   "DB302_HMI_Faults_Carrier71_Faults_1" : Int = PLC DB302_HMI_Faults.Carrier71_Faults_1 AT %DB1.DBW0, 1 s
   "DB302_HMI_Faults_Carrier71_Faults_2" : Int = PLC DB302_HMI_Faults.Carrier71_Faults_2 AT %DB1.DBW0, 1 s
   "DB302_HMI_Faults_Carrier71_Faults_3" : Int = PLC DB302_HMI_Faults.Carrier71_Faults_3 AT %DB1.DBW0, 1 s
   "DB302_HMI_Faults_Carrier72_Faults_0" : Int = PLC DB302_HMI_Faults.Carrier72_Faults_0 AT %DB1.DBW0, 1 s
   "DB302_HMI_Faults_Carrier72_Faults_1" : Int = PLC DB302_HMI_Faults.Carrier72_Faults_1 AT %DB1.DBW0, 1 s
   "DB302_HMI_Faults_Carrier72_Faults_2" : Int = PLC DB302_HMI_Faults.Carrier72_Faults_2 AT %DB1.DBW0, 1 s
   "DB302_HMI_Faults_Carrier72_Faults_3" : Int = PLC DB302_HMI_Faults.Carrier72_Faults_3 AT %DB1.DBW0, 1 s
   "DB302_HMI_Faults_Carrier73_Faults_0" : Int = PLC DB302_HMI_Faults.Carrier73_Faults_0 AT %DB1.DBW0, 1 s
   "DB302_HMI_Faults_Carrier73_Faults_1" : Int = PLC DB302_HMI_Faults.Carrier73_Faults_1 AT %DB1.DBW0, 1 s
   "DB302_HMI_Faults_Carrier73_Faults_2" : Int = PLC DB302_HMI_Faults.Carrier73_Faults_2 AT %DB1.DBW0, 1 s
   "DB302_HMI_Faults_Carrier73_Faults_3" : Int = PLC DB302_HMI_Faults.Carrier73_Faults_3 AT %DB1.DBW0, 1 s
   "DB302_HMI_Faults_Carrier74_Faults_0" : Int = PLC DB302_HMI_Faults.Carrier74_Faults_0 AT %DB1.DBW0, 1 s
   "DB302_HMI_Faults_Carrier74_Faults_1" : Int = PLC DB302_HMI_Faults.Carrier74_Faults_1 AT %DB1.DBW0, 1 s
   "DB302_HMI_Faults_Carrier74_Faults_2" : Int = PLC DB302_HMI_Faults.Carrier74_Faults_2 AT %DB1.DBW0, 1 s
   "DB302_HMI_Faults_Carrier74_Faults_3" : Int = PLC DB302_HMI_Faults.Carrier74_Faults_3 AT %DB1.DBW0, 1 s
   "DB302_HMI_Faults_Carrier75_Faults_0" : Int = PLC DB302_HMI_Faults.Carrier75_Faults_0 AT %DB1.DBW0, 1 s
   "DB302_HMI_Faults_Carrier75_Faults_1" : Int = PLC DB302_HMI_Faults.Carrier75_Faults_1 AT %DB1.DBW0, 1 s
   "DB302_HMI_Faults_Carrier75_Faults_2" : Int = PLC DB302_HMI_Faults.Carrier75_Faults_2 AT %DB1.DBW0, 1 s
   "DB302_HMI_Faults_Carrier75_Faults_3" : Int = PLC DB302_HMI_Faults.Carrier75_Faults_3 AT %DB1.DBW0, 1 s
   "DB302_HMI_Faults_Carrier76_Faults_0" : Int = PLC DB302_HMI_Faults.Carrier76_Faults_0 AT %DB1.DBW0, 1 s
   "DB302_HMI_Faults_Carrier76_Faults_1" : Int = PLC DB302_HMI_Faults.Carrier76_Faults_1 AT %DB1.DBW0, 1 s
   "DB302_HMI_Faults_Carrier76_Faults_2" : Int = PLC DB302_HMI_Faults.Carrier76_Faults_2 AT %DB1.DBW0, 1 s
   "DB302_HMI_Faults_Carrier76_Faults_3" : Int = PLC DB302_HMI_Faults.Carrier76_Faults_3 AT %DB1.DBW0, 1 s
   "DB302_HMI_Faults_Carrier77_Faults_0" : Int = PLC DB302_HMI_Faults.Carrier77_Faults_0 AT %DB1.DBW0, 1 s
   "DB302_HMI_Faults_Carrier77_Faults_1" : Int = PLC DB302_HMI_Faults.Carrier77_Faults_1 AT %DB1.DBW0, 1 s
   "DB302_HMI_Faults_Carrier77_Faults_2" : Int = PLC DB302_HMI_Faults.Carrier77_Faults_2 AT %DB1.DBW0, 1 s
   "DB302_HMI_Faults_Carrier77_Faults_3" : Int = PLC DB302_HMI_Faults.Carrier77_Faults_3 AT %DB1.DBW0, 1 s
   "DB302_HMI_Faults_Carrier78_Faults_0" : Int = PLC DB302_HMI_Faults.Carrier78_Faults_0 AT %DB1.DBW0, 1 s
   "DB302_HMI_Faults_Carrier78_Faults_1" : Int = PLC DB302_HMI_Faults.Carrier78_Faults_1 AT %DB1.DBW0, 1 s
   "DB302_HMI_Faults_Carrier78_Faults_2" : Int = PLC DB302_HMI_Faults.Carrier78_Faults_2 AT %DB1.DBW0, 1 s
   "DB302_HMI_Faults_Carrier78_Faults_3" : Int = PLC DB302_HMI_Faults.Carrier78_Faults_3 AT %DB1.DBW0, 1 s
   "DB302_HMI_Faults_Carrier79_Faults_0" : Int = PLC DB302_HMI_Faults.Carrier79_Faults_0 AT %DB1.DBW0, 1 s
   "DB302_HMI_Faults_Carrier79_Faults_1" : Int = PLC DB302_HMI_Faults.Carrier79_Faults_1 AT %DB1.DBW0, 1 s
   "DB302_HMI_Faults_Carrier79_Faults_2" : Int = PLC DB302_HMI_Faults.Carrier79_Faults_2 AT %DB1.DBW0, 1 s
   "DB302_HMI_Faults_Carrier79_Faults_3" : Int = PLC DB302_HMI_Faults.Carrier79_Faults_3 AT %DB1.DBW0, 1 s
   "DB302_HMI_Faults_Carrier8_Faults_0" : Int = PLC DB302_HMI_Faults.Carrier8_Faults_0 AT %DB1.DBW0, 1 s
   "DB302_HMI_Faults_Carrier8_Faults_1" : Int = PLC DB302_HMI_Faults.Carrier8_Faults_1 AT %DB1.DBW0, 1 s
   "DB302_HMI_Faults_Carrier8_Faults_2" : Int = PLC DB302_HMI_Faults.Carrier8_Faults_2 AT %DB1.DBW0, 1 s
   "DB302_HMI_Faults_Carrier8_Faults_3" : Int = PLC DB302_HMI_Faults.Carrier8_Faults_3 AT %DB1.DBW0, 1 s
   "DB302_HMI_Faults_Carrier80_Faults_0" : Int = PLC DB302_HMI_Faults.Carrier80_Faults_0 AT %DB1.DBW0, 1 s
   "DB302_HMI_Faults_Carrier80_Faults_1" : Int = PLC DB302_HMI_Faults.Carrier80_Faults_1 AT %DB1.DBW0, 1 s
   "DB302_HMI_Faults_Carrier80_Faults_2" : Int = PLC DB302_HMI_Faults.Carrier80_Faults_2 AT %DB1.DBW0, 1 s
   "DB302_HMI_Faults_Carrier80_Faults_3" : Int = PLC DB302_HMI_Faults.Carrier80_Faults_3 AT %DB1.DBW0, 1 s
   "DB302_HMI_Faults_Carrier81_Faults_0" : Int = PLC DB302_HMI_Faults.Carrier81_Faults_0 AT %DB1.DBW0, 1 s
   "DB302_HMI_Faults_Carrier81_Faults_1" : Int = PLC DB302_HMI_Faults.Carrier81_Faults_1 AT %DB1.DBW0, 1 s
   "DB302_HMI_Faults_Carrier81_Faults_2" : Int = PLC DB302_HMI_Faults.Carrier81_Faults_2 AT %DB1.DBW0, 1 s
   "DB302_HMI_Faults_Carrier81_Faults_3" : Int = PLC DB302_HMI_Faults.Carrier81_Faults_3 AT %DB1.DBW0, 1 s
   "DB302_HMI_Faults_Carrier82_Faults_0" : Int = PLC DB302_HMI_Faults.Carrier82_Faults_0 AT %DB1.DBW0, 1 s
   "DB302_HMI_Faults_Carrier82_Faults_1" : Int = PLC DB302_HMI_Faults.Carrier82_Faults_1 AT %DB1.DBW0, 1 s
   "DB302_HMI_Faults_Carrier82_Faults_2" : Int = PLC DB302_HMI_Faults.Carrier82_Faults_2 AT %DB1.DBW0, 1 s
   "DB302_HMI_Faults_Carrier82_Faults_3" : Int = PLC DB302_HMI_Faults.Carrier82_Faults_3 AT %DB1.DBW0, 1 s
   "DB302_HMI_Faults_Carrier9_Faults_0" : Int = PLC DB302_HMI_Faults.Carrier9_Faults_0 AT %DB1.DBW0, 1 s
   "DB302_HMI_Faults_Carrier9_Faults_1" : Int = PLC DB302_HMI_Faults.Carrier9_Faults_1 AT %DB1.DBW0, 1 s
   "DB302_HMI_Faults_Carrier9_Faults_2" : Int = PLC DB302_HMI_Faults.Carrier9_Faults_2 AT %DB1.DBW0, 1 s
   "DB302_HMI_Faults_Carrier9_Faults_3" : Int = PLC DB302_HMI_Faults.Carrier9_Faults_3 AT %DB1.DBW0, 1 s
   "DB401_HMI_Status_ZoneStatus.AccumZoneSpacing" : Word = PLC DB401_HMI_Status.ZoneStatus.AccumZoneSpacing, 1 s
   "DB401_HMI_Status_ZoneStatus.NextZoneNumber" : Int = PLC DB401_HMI_Status.ZoneStatus.NextZoneNumber, 1 s
   "DB401_HMI_Status_ZoneStatus.ProductionZoneSpacing" : Word = PLC DB401_HMI_Status.ZoneStatus.ProductionZoneSpacing, 1 s
   "DB401_HMI_Status_ZoneStatus.SpeedZone" : Bool = PLC DB401_HMI_Status.ZoneStatus.SpeedZone, 1 s
   "DB401_HMI_Status_ZoneStatus.SpeedZoneEndPos" : DWord = PLC DB401_HMI_Status.ZoneStatus.SpeedZoneEndPos, 1 s
   "DB401_HMI_Status_ZoneStatus.SpeedZoneStartPos" : DWord = PLC DB401_HMI_Status.ZoneStatus.SpeedZoneStartPos, 1 s
   "DB401_HMI_Status_ZoneStatus.ZoneEndPosition" : DWord = PLC DB401_HMI_Status.ZoneStatus.ZoneEndPosition, 1 s
   "DB401_HMI_Status_ZoneStatus.ZoneFull" : Bool = PLC DB401_HMI_Status.ZoneStatus.ZoneFull, 1 s
   "DB401_HMI_Status_ZoneStatus.ZoneIndex" : Int = PLC DB401_HMI_Status.ZoneStatus.ZoneIndex, 1 s
   "DB401_HMI_Status_ZoneStatus.ZoneStartPosition" : DWord = PLC DB401_HMI_Status.ZoneStatus.ZoneStartPosition, 1 s
   "DB401_HMI_Status_ZoneStatus.ZoneType" : String[254] = PLC DB401_HMI_Status.ZoneStatus.ZoneType, 1 s
   "DB401_HMI_Status_CarrierFaultCode" : Int = PLC DB401_HMI_Status.Status.CarrierFaultCode, 1 s
   "EMS_Zone[31]" : UDT_ZoneStructure = PLC EMS.Zone[31] AT %DB8.DBX31020.0, 1 s
   "EMS_Zone[32]" : UDT_ZoneStructure = PLC EMS.Zone[32] AT %DB8.DBX31020.0, 1 s
   "EMS_Zone[33]" : UDT_ZoneStructure = PLC EMS.Zone[33] AT %DB1.DBW0, 1 s
   "EMS_Zone[34]" : UDT_ZoneStructure = PLC EMS.Zone[34] AT %DB1.DBW0, 1 s
   "EMS_Zone[35]" : UDT_ZoneStructure = PLC EMS.Zone[35] AT %DB1.DBW0, 1 s
   "EMS_Zone[36]" : UDT_ZoneStructure = PLC EMS.Zone[36] AT %DB1.DBW0, 1 s
   "EMS_Zone[37]" : UDT_ZoneStructure = PLC EMS.Zone[37] AT %DB1.DBW0, 1 s
   "EMS_Zone[38]" : UDT_ZoneStructure = PLC EMS.Zone[38] AT %DB1.DBW0, 1 s
   "EMS_Zone[39]" : UDT_ZoneStructure = PLC EMS.Zone[39] AT %DB1.DBW0, 1 s
   "EMS_Zone[4]" : UDT_ZoneStructure = PLC EMS.Zone[4] AT %DB8.DBX4136.0, 1 s
   "EMS_Zone[40]" : UDT_ZoneStructure = PLC EMS.Zone[40] AT %DB1.DBW0, 1 s
   "EMS_Zone[41]" : UDT_ZoneStructure = PLC EMS.Zone[41] AT %DB1.DBW0, 1 s
   "EMS_Zone[42]" : UDT_ZoneStructure = PLC EMS.Zone[42] AT %DB1.DBW0, 1 s
   "EMS_Zone[43]" : UDT_ZoneStructure = PLC EMS.Zone[43] AT %DB1.DBW0, 1 s
   "EMS_Zone[44]" : UDT_ZoneStructure = PLC EMS.Zone[44] AT %DB1.DBW0, 1 s
   "EMS_Zone[45]" : UDT_ZoneStructure = PLC EMS.Zone[45] AT %DB1.DBW0, 1 s
   "EMS_Zone[46]" : UDT_ZoneStructure = PLC EMS.Zone[46] AT %DB1.DBW0, 1 s
   "EMS_Zone[47]" : UDT_ZoneStructure = PLC EMS.Zone[47] AT %DB1.DBW0, 1 s
   "EMS_Zone[48]" : UDT_ZoneStructure = PLC EMS.Zone[48] AT %DB1.DBW0, 1 s
   "EMS_Zone[49]" : UDT_ZoneStructure = PLC EMS.Zone[49] AT %DB1.DBW0, 1 s
   "EMS_Zone[5]" : UDT_ZoneStructure = PLC EMS.Zone[5] AT %DB8.DBX5170.0, 1 s
   "EMS_Zone[50]" : UDT_ZoneStructure = PLC EMS.Zone[50] AT %DB1.DBW0, 1 s
   "EMS_Zone[51]" : UDT_ZoneStructure = PLC EMS.Zone[51] AT %DB1.DBW0, 1 s
   "EMS_Zone[52]" : UDT_ZoneStructure = PLC EMS.Zone[52] AT %DB8.DBX31020.0, 1 s
   "EMS_Zone[53]" : UDT_ZoneStructure = PLC EMS.Zone[53] AT %DB1.DBW0, 1 s
   "EMS_Zone[54]" : UDT_ZoneStructure = PLC EMS.Zone[54] AT %DB1.DBW0, 1 s
   "EMS_Zone[55]" : UDT_ZoneStructure = PLC EMS.Zone[55] AT %DB1.DBW0, 1 s
   "EMS_Zone[56]" : UDT_ZoneStructure = PLC EMS.Zone[56] AT %DB1.DBW0, 1 s
   "EMS_Zone[57]" : UDT_ZoneStructure = PLC EMS.Zone[57] AT %DB1.DBW0, 1 s
   "EMS_Zone[58]" : UDT_ZoneStructure = PLC EMS.Zone[58] AT %DB8.DBX31020.0, 1 s
   "EMS_Zone[59]" : UDT_ZoneStructure = PLC EMS.Zone[59] AT %DB1.DBW0, 1 s
   "EMS_Zone[6]" : UDT_ZoneStructure = PLC EMS.Zone[6] AT %DB8.DBX6204.0, 1 s
   "EMS_Zone[60]" : UDT_ZoneStructure = PLC EMS.Zone[60] AT %DB1.DBW0, 1 s
   "EMS_Zone[61]" : UDT_ZoneStructure = PLC EMS.Zone[61] AT %DB1.DBW0, 1 s
   "EMS_Zone[62]" : UDT_ZoneStructure = PLC EMS.Zone[62] AT %DB1.DBW0, 1 s
   "EMS_Zone[63]" : UDT_ZoneStructure = PLC EMS.Zone[63] AT %DB1.DBW0, 1 s
   "DB401_HMI_Status_ZoneStatus.PrevZoneNumber" : Int = PLC DB401_HMI_Status.ZoneStatus.PrevZoneNumber, 1 s
   "Mask_Carrier_Faults_LT" : Bool = PLC DB401_HMI_Status.Status.MaskCarrierFaultsLT AT %DB1.DBX0.0, 1 s
   "Reset_Mask_Carrier_Faults_PB" : Bool = PLC DB401_HMI_Status.Status.ResetMaskCarrierFaultsPB AT %DB1.DBX0.0, 1 s
   "Set_Mask_Carrier_Faults_PB" : Bool = PLC DB401_HMI_Status.Status.SetMaskCarrierFaultsPB AT %DB1.DBX0.0, 1 s
   "HMI_Carrier_CurrentArea" : String[2] = PLC DB401_HMI_Status.Status.Area AT %DB1.DBW0, 1 s

HMI tags "SDC"
   "Clock_1Hz" : Bool = PLC Clock_1Hz AT %M0.5, 500 ms   // Zyklusflanke 1Hz / Cycle flag 1Hz
   "SDC\_EDIT" : Int, internal
   "SDC\_EDIT_BIT" : Bool, internal
   "SDC\_open_EMS_Stat" : Bool, internal
      on ChangeValue: ActivateScreen("711_CARRIER_STATUS", 0)
   "SDC\_open_Section_Para" : Bool, internal
      on ChangeValue: ActivateScreen("708_ZONE_STATUS", 0)
   "HMI_EMS_Nr" : Int = PLC HMI_EMS_Nr AT %MW30, 1 s
   "SDC\_TS_Nr" : Int, internal
      on ChangeValue: "SDC_TS_PARAMETER"(); "SDC_TS_REFERENCE"("SDC\_TS_Nr")
   "SDC\_intern_Bildnummer" : Int AT %DB1.DBX0.0
   "DB_SDC_GLOBAL_M.SDC_ER_Reset" : Bool = PLC DB_SDC_GLOBAL.M.SDC_ER_Reset AT %DB3700.DBX600.4, 1 s
   "SDC\_intern_MELDUNGEN" : Int, internal
   "SDC\_Pos_sichtbar" : Bool AT %DB1.DBX4.0
   "AlwaysTRUE" : Bool = PLC AlwaysTRUE AT %M1.2, 500 ms
   "AlwaysFALSE" : Bool = PLC AlwaysFALSE AT %M1.3, 500 ms
   "HMI_Zone_Nr" : Int = PLC HMI_Zone_Nr AT %MW102, 1 s
   "HMI_Status_G120D_Control" : Word = PLC DB401_HMI_Status.Drive.G120D_CONTROL AT %DB1.DBW0, 1 s
   "HMI_Status_G120D_Status" : Word = PLC DB401_HMI_Status.Drive.G120D_STATUS AT %DB1.DBW0, 1 s
   "HMI_Status_Slot2_Inputs" : Byte = PLC DB401_HMI_Status.IO.Carrier_Slot02_Inputs AT %DB1.DBW0, 1 s
   "HMI_Status_Slot3_Outputs" : Byte = PLC DB401_HMI_Status.IO.Carrier_Slot03_Outputs AT %DB1.DBW0, 1 s
   "HMI_Status_Slot4_Inputs" : Word = PLC DB401_HMI_Status.IO.Carrier_Slot04_Inputs AT %DB1.DBW0, 1 s
   "HMI_Status_Slot5_Outputs" : Word = PLC DB401_HMI_Status.IO.Carrier_Slot05_Outputs AT %DB1.DBW0, 1 s
   "HMI_Carrier_Comm_Fault" : Bool = PLC DB401_HMI_Status.Status.CommFlt AT %DB1.DBW0, 1 s
   "HMI_Carrier_Faulted" : Bool = PLC DB401_HMI_Status.Status.Faulted AT %DB1.DBW0, 1 s
   "HMI_Carrier_Auto" : Bool = PLC DB401_HMI_Status.Status.AutoMode AT %DB1.DBW0, 1 s
   "HMI_Carrier_Manual" : Bool = PLC DB401_HMI_Status.Status.ManualMode AT %DB1.DBW0, 1 s
   "HMI_Carrier_RunningFwd" : Bool = PLC DB401_HMI_Status.Status.RunningFWD AT %DB1.DBW0, 1 s
   "HMI_Carrier_RunningRev" : Bool = PLC DB401_HMI_Status.Status.RunningREV AT %DB1.DBW0, 1 s
   "HMI_Carrier_HoldPBPressed" : Bool = PLC DB401_HMI_Status.Status.ProductionHoldPB_Status AT %DB1.DBW0, 1 s
   "HMI_Carrier_DriveFwdCommand" : Bool = PLC DB401_HMI_Status.Status.DriveFwdCMD AT %DB1.DBW0, 1 s
   "HMI_Carrier_DriveCmdSpeed" : Word = PLC DB401_HMI_Status.Status.DriveCmdSpeed AT %DB1.DBW0, 1 s
   "HMI_Carrier_CurrentPosition" : DWord = PLC DB401_HMI_Status.Status.CarrierPosition AT %DB1.DBW0, 1 s
   "HMI_Carrier_ActualSpeed" : Word = PLC DB401_HMI_Status.Status.ActualSpeed AT %DB1.DBW0, 1 s
   "HMI_Carrier_NextCarrierNumber" : Word = PLC DB401_HMI_Status.Status.NextCarrierNum AT %DB1.DBW0, 1 s
   "HMI_Carrier_CurrentZone" : Int = PLC DB401_HMI_Status.Status.Zone AT %DB1.DBW0, 1 s
   "HMI_Carrier_AtCommandPosition" : Bool = PLC DB401_HMI_Status.Status.AtCmdPos AT %DB1.DBW0, 1 s
   "HMI_Carrier_NextStopPosition" : DWord = PLC DB401_HMI_Status.Status.NextStopPosition AT %DB1.DBW0, 1 s
   "HMI_Carrier_DriveCommFault" : Bool = PLC DB401_HMI_Status.Status.DriveCommFault AT %DB1.DBW0, 1 s
   "HMI_Carrier_EncoderCommFault" : Bool = PLC DB401_HMI_Status.Status.EncoderCommFault AT %DB1.DBW0, 1 s
   "HMI_Carrier_HMICommFault" : Bool = PLC DB401_HMI_Status.Status.HMICommFault AT %DB1.DBW0, 1 s

HMI tags "DB_SDC_EMS_TS_HMI"
   "DB_SDC_EMS_TS_1_HMI_SEK[88].EMS[1]" : UDT_SDC_EMS_TS_STAT_HMI = PLC DB_SDC_EMS_TS_1_HMI.SEK[88].EMS[1] AT %DB3810.DBX15680.0, 1 s
   "DB_SDC_EMS_TS_1_HMI_SEK[89].EMS[1]" : UDT_SDC_EMS_TS_STAT_HMI = PLC DB_SDC_EMS_TS_1_HMI.SEK[89].EMS[1] AT %DB3810.DBX15860.0, 1 s
   "DB_SDC_EMS_TS_1_HMI_SEK[90].EMS[1]" : UDT_SDC_EMS_TS_STAT_HMI = PLC DB_SDC_EMS_TS_1_HMI.SEK[90].EMS[1] AT %DB3810.DBX16040.0, 1 s
   "DB_SDC_EMS_TS_1_HMI_SEK[91].EMS[1]" : UDT_SDC_EMS_TS_STAT_HMI = PLC DB_SDC_EMS_TS_1_HMI.SEK[91].EMS[1] AT %DB3810.DBX16220.0, 1 s
   "DB_SDC_EMS_TS_1_HMI_SEK[92].EMS[1]" : UDT_SDC_EMS_TS_STAT_HMI = PLC DB_SDC_EMS_TS_1_HMI.SEK[92].EMS[1] AT %DB3810.DBX16400.0, 1 s
   "DB_SDC_EMS_TS_1_HMI_SEK[93].EMS[1]" : UDT_SDC_EMS_TS_STAT_HMI = PLC DB_SDC_EMS_TS_1_HMI.SEK[93].EMS[1] AT %DB3810.DBX16580.0, 1 s
   "DB_SDC_EMS_TS_1_HMI_SEK[94].EMS[1]" : UDT_SDC_EMS_TS_STAT_HMI = PLC DB_SDC_EMS_TS_1_HMI.SEK[94].EMS[1] AT %DB3810.DBX16760.0, 1 s
   "DB_SDC_EMS_TS_1_HMI_SEK[95].EMS[1]" : UDT_SDC_EMS_TS_STAT_HMI = PLC DB_SDC_EMS_TS_1_HMI.SEK[95].EMS[1] AT %DB3810.DBX16940.0, 1 s
   "DB_SDC_EMS_TS_1_HMI_SEK[96].EMS[1]" : UDT_SDC_EMS_TS_STAT_HMI = PLC DB_SDC_EMS_TS_1_HMI.SEK[96].EMS[1] AT %DB3810.DBX17120.0, 1 s
   "DB_SDC_EMS_TS_1_HMI_SEK[100].EMS[1]" : UDT_SDC_EMS_TS_STAT_HMI = PLC DB_SDC_EMS_TS_1_HMI.SEK[100].EMS[1] AT %DB3810.DBX17840.0, 1 s
   "DB_SDC_EMS_TS_1_HMI_SEK[101].EMS[1]" : UDT_SDC_EMS_TS_STAT_HMI = PLC DB_SDC_EMS_TS_1_HMI.SEK[101].EMS[1] AT %DB3810.DBX18020.0, 1 s
   "DB_SDC_EMS_TS_1_HMI_SEK[102].EMS[1]" : UDT_SDC_EMS_TS_STAT_HMI = PLC DB_SDC_EMS_TS_1_HMI.SEK[102].EMS[1] AT %DB3810.DBX18200.0, 1 s
   "DB_SDC_EMS_TS_1_HMI_SEK[103].EMS[1]" : UDT_SDC_EMS_TS_STAT_HMI = PLC DB_SDC_EMS_TS_1_HMI.SEK[103].EMS[1] AT %DB3810.DBX18380.0, 1 s
   "DB_SDC_EMS_TS_1_HMI_SEK[104].EMS[1]" : UDT_SDC_EMS_TS_STAT_HMI = PLC DB_SDC_EMS_TS_1_HMI.SEK[104].EMS[1] AT %DB3810.DBX18560.0, 1 s
   "DB_SDC_EMS_TS_1_HMI_SEK[105].EMS[1]" : UDT_SDC_EMS_TS_STAT_HMI = PLC DB_SDC_EMS_TS_1_HMI.SEK[105].EMS[1] AT %DB3810.DBX18740.0, 1 s
   "DB_SDC_EMS_TS_1_HMI_SEK[106].EMS[1]" : UDT_SDC_EMS_TS_STAT_HMI = PLC DB_SDC_EMS_TS_1_HMI.SEK[106].EMS[1] AT %DB3810.DBX18920.0, 1 s
   "DB_SDC_EMS_TS_1_HMI_SEK[107].EMS[1]" : UDT_SDC_EMS_TS_STAT_HMI = PLC DB_SDC_EMS_TS_1_HMI.SEK[107].EMS[1] AT %DB3810.DBX19100.0, 1 s
   "DB_SDC_EMS_TS_1_HMI_SEK[108].EMS[1]" : UDT_SDC_EMS_TS_STAT_HMI = PLC DB_SDC_EMS_TS_1_HMI.SEK[108].EMS[1] AT %DB3810.DBX19280.0, 1 s
   "DB_SDC_EMS_TS_1_HMI_SEK[109].EMS[1]" : UDT_SDC_EMS_TS_STAT_HMI = PLC DB_SDC_EMS_TS_1_HMI.SEK[109].EMS[1] AT %DB3810.DBX19460.0, 1 s
   "DB_SDC_EMS_TS_1_HMI_SEK[110].EMS[1]" : UDT_SDC_EMS_TS_STAT_HMI = PLC DB_SDC_EMS_TS_1_HMI.SEK[110].EMS[1] AT %DB3810.DBX19640.0, 1 s
   "DB_SDC_EMS_TS_1_HMI_SEK[111].EMS[1]" : UDT_SDC_EMS_TS_STAT_HMI = PLC DB_SDC_EMS_TS_1_HMI.SEK[111].EMS[1] AT %DB3810.DBX19820.0, 1 s
   "DB_SDC_EMS_TS_1_HMI_SEK[120].EMS[1]" : UDT_SDC_EMS_TS_STAT_HMI = PLC DB_SDC_EMS_TS_1_HMI.SEK[120].EMS[1] AT %DB3810.DBX21440.0, 1 s
   "DB_SDC_EMS_TS_1_HMI_SEK[121].EMS[1]" : UDT_SDC_EMS_TS_STAT_HMI = PLC DB_SDC_EMS_TS_1_HMI.SEK[121].EMS[1] AT %DB3810.DBX21620.0, 1 s
   "DB_SDC_EMS_TS_1_HMI_SEK[126].EMS[1]" : UDT_SDC_EMS_TS_STAT_HMI = PLC DB_SDC_EMS_TS_1_HMI.SEK[126].EMS[1] AT %DB3810.DBX22520.0, 1 s
   "DB_SDC_EMS_TS_1_HMI_SEK[125].EMS[1]" : UDT_SDC_EMS_TS_STAT_HMI = PLC DB_SDC_EMS_TS_1_HMI.SEK[125].EMS[1] AT %DB3810.DBX22340.0, 1 s
   "DB_SDC_EMS_TS_1_HMI_SEK[122].EMS[1]" : UDT_SDC_EMS_TS_STAT_HMI = PLC DB_SDC_EMS_TS_1_HMI.SEK[122].EMS[1] AT %DB3810.DBX21800.0, 1 s
   "DB_SDC_EMS_TS_1_HMI_SEK[123].EMS[1]" : UDT_SDC_EMS_TS_STAT_HMI = PLC DB_SDC_EMS_TS_1_HMI.SEK[123].EMS[1] AT %DB3810.DBX21980.0, 1 s
   "DB_SDC_EMS_TS_1_HMI_SEK[124].EMS[1]" : UDT_SDC_EMS_TS_STAT_HMI = PLC DB_SDC_EMS_TS_1_HMI.SEK[124].EMS[1] AT %DB3810.DBX22160.0, 1 s
   "DB_SDC_EMS_TS_1_HMI_SEK[127].EMS[1]" : UDT_SDC_EMS_TS_STAT_HMI = PLC DB_SDC_EMS_TS_1_HMI.SEK[127].EMS[1] AT %DB3810.DBX22700.0, 1 s
   "DB_SDC_EMS_TS_1_HMI_SEK[128].EMS[1]" : UDT_SDC_EMS_TS_STAT_HMI = PLC DB_SDC_EMS_TS_1_HMI.SEK[128].EMS[1] AT %DB3810.DBX22880.0, 1 s
   "DB_SDC_EMS_TS_1_HMI_SEK[129].EMS[1]" : UDT_SDC_EMS_TS_STAT_HMI = PLC DB_SDC_EMS_TS_1_HMI.SEK[129].EMS[1] AT %DB3810.DBX23060.0, 1 s
   "DB_SDC_EMS_TS_1_HMI_SEK[130].EMS[1]" : UDT_SDC_EMS_TS_STAT_HMI = PLC DB_SDC_EMS_TS_1_HMI.SEK[130].EMS[1] AT %DB3810.DBX23240.0, 1 s
   "DB_SDC_EMS_TS_1_HMI_SEK[131].EMS[1]" : UDT_SDC_EMS_TS_STAT_HMI = PLC DB_SDC_EMS_TS_1_HMI.SEK[131].EMS[1] AT %DB3810.DBX23420.0, 1 s
   "DB_SDC_EMS_TS_1_HMI_SEK[132].EMS[1]" : UDT_SDC_EMS_TS_STAT_HMI = PLC DB_SDC_EMS_TS_1_HMI.SEK[132].EMS[1] AT %DB3810.DBX23600.0, 1 s
   "DB_SDC_EMS_TS_1_HMI_SEK[140].EMS[1]" : UDT_SDC_EMS_TS_STAT_HMI = PLC DB_SDC_EMS_TS_1_HMI.SEK[140].EMS[1] AT %DB3810.DBX25040.0, 1 s
   "DB_SDC_EMS_TS_1_HMI_SEK[141].EMS[1]" : UDT_SDC_EMS_TS_STAT_HMI = PLC DB_SDC_EMS_TS_1_HMI.SEK[141].EMS[1] AT %DB3810.DBX25220.0, 1 s
   "DB_SDC_EMS_TS_1_HMI_SEK[142].EMS[1]" : UDT_SDC_EMS_TS_STAT_HMI = PLC DB_SDC_EMS_TS_1_HMI.SEK[142].EMS[1] AT %DB3810.DBX25400.0, 1 s
   "DB_SDC_EMS_TS_1_HMI_SEK[143].EMS[1]" : UDT_SDC_EMS_TS_STAT_HMI = PLC DB_SDC_EMS_TS_1_HMI.SEK[143].EMS[1] AT %DB3810.DBX25580.0, 1 s
   "DB_SDC_EMS_TS_1_HMI_SEK[144].EMS[1]" : UDT_SDC_EMS_TS_STAT_HMI = PLC DB_SDC_EMS_TS_1_HMI.SEK[144].EMS[1] AT %DB3810.DBX25760.0, 1 s
   "DB_SDC_EMS_TS_1_HMI_SEK[145].EMS[1]" : UDT_SDC_EMS_TS_STAT_HMI = PLC DB_SDC_EMS_TS_1_HMI.SEK[145].EMS[1] AT %DB3810.DBX25940.0, 1 s
   "DB_SDC_EMS_TS_1_HMI_SEK[146].EMS[1]" : UDT_SDC_EMS_TS_STAT_HMI = PLC DB_SDC_EMS_TS_1_HMI.SEK[146].EMS[1] AT %DB3810.DBX26120.0, 1 s
   "DB_SDC_EMS_TS_1_HMI_SEK[147].EMS[1]" : UDT_SDC_EMS_TS_STAT_HMI = PLC DB_SDC_EMS_TS_1_HMI.SEK[147].EMS[1] AT %DB3810.DBX26300.0, 1 s
   "DB_SDC_EMS_TS_1_HMI_SEK[148].EMS[1]" : UDT_SDC_EMS_TS_STAT_HMI = PLC DB_SDC_EMS_TS_1_HMI.SEK[148].EMS[1] AT %DB3810.DBX26480.0, 1 s
   "DB_SDC_EMS_TS_1_HMI_SEK[149].EMS[1]" : UDT_SDC_EMS_TS_STAT_HMI = PLC DB_SDC_EMS_TS_1_HMI.SEK[149].EMS[1] AT %DB3810.DBX26660.0, 1 s
   "DB_SDC_EMS_TS_1_HMI_SEK[150].EMS[1]" : UDT_SDC_EMS_TS_STAT_HMI = PLC DB_SDC_EMS_TS_1_HMI.SEK[150].EMS[1] AT %DB3810.DBX26840.0, 1 s
   "DB_SDC_EMS_TS_1_HMI_SEK[151].EMS[1]" : UDT_SDC_EMS_TS_STAT_HMI = PLC DB_SDC_EMS_TS_1_HMI.SEK[151].EMS[1] AT %DB3810.DBX27020.0, 1 s
   "DB_SDC_EMS_TS_1_HMI_SEK[152].EMS[1]" : UDT_SDC_EMS_TS_STAT_HMI = PLC DB_SDC_EMS_TS_1_HMI.SEK[152].EMS[1] AT %DB3810.DBX27200.0, 1 s
   "DB_SDC_EMS_TS_1_HMI_SEK[160].EMS[1]" : UDT_SDC_EMS_TS_STAT_HMI = PLC DB_SDC_EMS_TS_1_HMI.SEK[160].EMS[1] AT %DB3810.DBX28640.0, 1 s
   "DB_SDC_EMS_TS_1_HMI_SEK[161].EMS[1]" : UDT_SDC_EMS_TS_STAT_HMI = PLC DB_SDC_EMS_TS_1_HMI.SEK[161].EMS[1] AT %DB3810.DBX28820.0, 1 s
   "DB_SDC_EMS_TS_1_HMI_SEK[162].EMS[1]" : UDT_SDC_EMS_TS_STAT_HMI = PLC DB_SDC_EMS_TS_1_HMI.SEK[162].EMS[1] AT %DB3810.DBX29000.0, 1 s
   "DB_SDC_EMS_TS_1_HMI_SEK[163].EMS[1]" : UDT_SDC_EMS_TS_STAT_HMI = PLC DB_SDC_EMS_TS_1_HMI.SEK[163].EMS[1] AT %DB3810.DBX29180.0, 1 s
   "DB_SDC_EMS_TS_1_HMI_SEK[164].EMS[1]" : UDT_SDC_EMS_TS_STAT_HMI = PLC DB_SDC_EMS_TS_1_HMI.SEK[164].EMS[1] AT %DB3810.DBX29360.0, 1 s
   "DB_SDC_EMS_TS_1_HMI_SEK[165].EMS[1]" : UDT_SDC_EMS_TS_STAT_HMI = PLC DB_SDC_EMS_TS_1_HMI.SEK[165].EMS[1] AT %DB3810.DBX29540.0, 1 s
   "DB_SDC_EMS_TS_1_HMI_SEK[166].EMS[1]" : UDT_SDC_EMS_TS_STAT_HMI = PLC DB_SDC_EMS_TS_1_HMI.SEK[166].EMS[1] AT %DB3810.DBX29720.0, 1 s
   "DB_SDC_EMS_TS_1_HMI_SEK[167].EMS[1]" : UDT_SDC_EMS_TS_STAT_HMI = PLC DB_SDC_EMS_TS_1_HMI.SEK[167].EMS[1] AT %DB3810.DBX29900.0, 1 s
   "DB_SDC_EMS_TS_1_HMI_SEK[168].EMS[1]" : UDT_SDC_EMS_TS_STAT_HMI = PLC DB_SDC_EMS_TS_1_HMI.SEK[168].EMS[1] AT %DB3810.DBX30080.0, 1 s
   "DB_SDC_EMS_TS_1_HMI_SEK[169].EMS[1]" : UDT_SDC_EMS_TS_STAT_HMI = PLC DB_SDC_EMS_TS_1_HMI.SEK[169].EMS[1] AT %DB3810.DBX30260.0, 1 s
   "DB_SDC_EMS_TS_1_HMI_SEK[170].EMS[1]" : UDT_SDC_EMS_TS_STAT_HMI = PLC DB_SDC_EMS_TS_1_HMI.SEK[170].EMS[1] AT %DB3810.DBX30440.0, 1 s
   "DB_SDC_EMS_TS_1_HMI_SEK[190].EMS[1]" : UDT_SDC_EMS_TS_STAT_HMI = PLC DB_SDC_EMS_TS_1_HMI.SEK[190].EMS[1] AT %DB3810.DBX34040.0, 1 s
   "DB_SDC_EMS_TS_1_HMI_SEK[191].EMS[1]" : UDT_SDC_EMS_TS_STAT_HMI = PLC DB_SDC_EMS_TS_1_HMI.SEK[191].EMS[1] AT %DB3810.DBX34220.0, 1 s
   "DB_SDC_EMS_TS_1_HMI_SEK[192].EMS[1]" : UDT_SDC_EMS_TS_STAT_HMI = PLC DB_SDC_EMS_TS_1_HMI.SEK[192].EMS[1] AT %DB3810.DBX34400.0, 1 s
   "DB_SDC_EMS_TS_1_HMI_SEK[193].EMS[1]" : UDT_SDC_EMS_TS_STAT_HMI = PLC DB_SDC_EMS_TS_1_HMI.SEK[193].EMS[1] AT %DB3810.DBX34580.0, 1 s
   "DB_SDC_EMS_TS_1_HMI_SEK[194].EMS[1]" : UDT_SDC_EMS_TS_STAT_HMI = PLC DB_SDC_EMS_TS_1_HMI.SEK[194].EMS[1] AT %DB3810.DBX34760.0, 1 s
   "DB_SDC_EMS_TS_1_HMI_SEK[195].EMS[1]" : UDT_SDC_EMS_TS_STAT_HMI = PLC DB_SDC_EMS_TS_1_HMI.SEK[195].EMS[1] AT %DB3810.DBX34940.0, 1 s
   "DB_SDC_EMS_TS_1_HMI_SEK[86].EMS[1]" : UDT_SDC_EMS_TS_STAT_HMI = PLC DB_SDC_EMS_TS_1_HMI.SEK[86].EMS[1] AT %DB3810.DBX15320.0, 1 s
   "DB_SDC_EMS_TS_1_HMI_SEK[87].EMS[1]" : UDT_SDC_EMS_TS_STAT_HMI = PLC DB_SDC_EMS_TS_1_HMI.SEK[87].EMS[1] AT %DB3810.DBX15500.0, 1 s
   "DB_SDC_EMS_TS_1_HMI_SEK[137].EMS[1]" : UDT_SDC_EMS_TS_STAT_HMI = PLC DB_SDC_EMS_TS_1_HMI.SEK[137].EMS[1] AT %DB3810.DBX24500.0, 1 s
   "DB_SDC_EMS_TS_1_HMI_SEK[136].EMS[1]" : UDT_SDC_EMS_TS_STAT_HMI = PLC DB_SDC_EMS_TS_1_HMI.SEK[136].EMS[1] AT %DB3810.DBX24320.0, 1 s
   "DB_SDC_EMS_TS_1_HMI_SEK[135].EMS[1]" : UDT_SDC_EMS_TS_STAT_HMI = PLC DB_SDC_EMS_TS_1_HMI.SEK[135].EMS[1] AT %DB3810.DBX24140.0, 1 s
   "DB_SDC_EMS_TS_1_HMI_SEK[134].EMS[1]" : UDT_SDC_EMS_TS_STAT_HMI = PLC DB_SDC_EMS_TS_1_HMI.SEK[134].EMS[1] AT %DB3810.DBX23960.0, 1 s

HMI tags "DB_SDC_EMS_TS_HMI_BA2"
   "DB_SDC_EMS_TS_1_HMI_SEK[99].EMS[1]" : UDT_SDC_EMS_TS_STAT_HMI = PLC DB_SDC_EMS_TS_1_HMI.SEK[99].EMS[1] AT %DB3810.DBX17660.0, 1 s
   "DB_SDC_EMS_TS_1_HMI_SEK[100].EMS[1](1)" : UDT_SDC_EMS_TS_STAT_HMI = PLC DB_SDC_EMS_TS_1_HMI.SEK[100].EMS[1] AT %DB3810.DBX17840.0, 1 s
   "DB_SDC_EMS_TS_1_HMI_SEK[101].EMS[1](1)" : UDT_SDC_EMS_TS_STAT_HMI = PLC DB_SDC_EMS_TS_1_HMI.SEK[101].EMS[1] AT %DB3810.DBX18020.0, 1 s
   "DB_SDC_EMS_TS_1_HMI_SEK[102].EMS[1](1)" : UDT_SDC_EMS_TS_STAT_HMI = PLC DB_SDC_EMS_TS_1_HMI.SEK[102].EMS[1] AT %DB3810.DBX18200.0, 1 s
   "DB_SDC_EMS_TS_1_HMI_SEK[103].EMS[1](1)" : UDT_SDC_EMS_TS_STAT_HMI = PLC DB_SDC_EMS_TS_1_HMI.SEK[103].EMS[1] AT %DB3810.DBX18380.0, 1 s
   "DB_SDC_EMS_TS_1_HMI_SEK[104].EMS[1](1)" : UDT_SDC_EMS_TS_STAT_HMI = PLC DB_SDC_EMS_TS_1_HMI.SEK[104].EMS[1] AT %DB3810.DBX18560.0, 1 s
   "DB_SDC_EMS_TS_1_HMI_SEK[105].EMS[1](1)" : UDT_SDC_EMS_TS_STAT_HMI = PLC DB_SDC_EMS_TS_1_HMI.SEK[105].EMS[1] AT %DB3810.DBX18740.0, 1 s
   "DB_SDC_EMS_TS_1_HMI_SEK[106].EMS[1](1)" : UDT_SDC_EMS_TS_STAT_HMI = PLC DB_SDC_EMS_TS_1_HMI.SEK[106].EMS[1] AT %DB3810.DBX18920.0, 1 s
   "DB_SDC_EMS_TS_1_HMI_SEK[107].EMS[1](1)" : UDT_SDC_EMS_TS_STAT_HMI = PLC DB_SDC_EMS_TS_1_HMI.SEK[107].EMS[1] AT %DB3810.DBX19100.0, 1 s
   "DB_SDC_EMS_TS_1_HMI_SEK[108].EMS[1](1)" : UDT_SDC_EMS_TS_STAT_HMI = PLC DB_SDC_EMS_TS_1_HMI.SEK[108].EMS[1] AT %DB3810.DBX19280.0, 1 s
   "DB_SDC_EMS_TS_1_HMI_SEK[109].EMS[1](1)" : UDT_SDC_EMS_TS_STAT_HMI = PLC DB_SDC_EMS_TS_1_HMI.SEK[109].EMS[1] AT %DB3810.DBX19460.0, 1 s
   "DB_SDC_EMS_TS_1_HMI_SEK[110].EMS[1](1)" : UDT_SDC_EMS_TS_STAT_HMI = PLC DB_SDC_EMS_TS_1_HMI.SEK[110].EMS[1] AT %DB3810.DBX19640.0, 1 s
   "DB_SDC_EMS_TS_1_HMI_SEK[111].EMS[1](1)" : UDT_SDC_EMS_TS_STAT_HMI = PLC DB_SDC_EMS_TS_1_HMI.SEK[111].EMS[1] AT %DB3810.DBX19820.0, 1 s
   "DB_SDC_EMS_TS_1_HMI_SEK[112].EMS[1]" : UDT_SDC_EMS_TS_STAT_HMI = PLC DB_SDC_EMS_TS_1_HMI.SEK[112].EMS[1] AT %DB3810.DBX20000.0, 1 s
   "DB_SDC_EMS_TS_1_HMI_SEK[113].EMS[1]" : UDT_SDC_EMS_TS_STAT_HMI = PLC DB_SDC_EMS_TS_1_HMI.SEK[113].EMS[1] AT %DB3810.DBX20180.0, 1 s
   "DB_SDC_EMS_TS_1_HMI_SEK[114].EMS[1]" : UDT_SDC_EMS_TS_STAT_HMI = PLC DB_SDC_EMS_TS_1_HMI.SEK[114].EMS[1] AT %DB3810.DBX20360.0, 1 s
   "DB_SDC_EMS_TS_1_HMI_SEK[99].EMS[2]" : UDT_SDC_EMS_TS_STAT_HMI = PLC DB_SDC_EMS_TS_1_HMI.SEK[99].EMS[2] AT %DB3810.DBX17690.0, 1 s
   "DB_SDC_EMS_TS_1_HMI_SEK[100].EMS[2]" : UDT_SDC_EMS_TS_STAT_HMI = PLC DB_SDC_EMS_TS_1_HMI.SEK[100].EMS[2] AT %DB3810.DBX17870.0, 1 s
   "DB_SDC_EMS_TS_1_HMI_SEK[2]" : UDT_SDC_6EMS_TS_STAT_HMI = PLC DB_SDC_EMS_TS_1_HMI.SEK[2] AT %DB3810.DBX200.0, 1 s
   "DB_SDC_EMS_TS_1_HMI_SEK[102].EMS[2]" : UDT_SDC_EMS_TS_STAT_HMI = PLC DB_SDC_EMS_TS_1_HMI.SEK[102].EMS[2] AT %DB3810.DBX18230.0, 1 s
   "DB_SDC_EMS_TS_1_HMI_SEK[103].EMS[2]" : UDT_SDC_EMS_TS_STAT_HMI = PLC DB_SDC_EMS_TS_1_HMI.SEK[103].EMS[2] AT %DB3810.DBX18410.0, 1 s
   "DB_SDC_EMS_TS_1_HMI_SEK[104].EMS[2]" : UDT_SDC_EMS_TS_STAT_HMI = PLC DB_SDC_EMS_TS_1_HMI.SEK[104].EMS[2] AT %DB3810.DBX18590.0, 1 s
   "DB_SDC_EMS_TS_1_HMI_SEK[105].EMS[2]" : UDT_SDC_EMS_TS_STAT_HMI = PLC DB_SDC_EMS_TS_1_HMI.SEK[105].EMS[2] AT %DB3810.DBX18770.0, 1 s
   "DB_SDC_EMS_TS_1_HMI_SEK[106].EMS[2]" : UDT_SDC_EMS_TS_STAT_HMI = PLC DB_SDC_EMS_TS_1_HMI.SEK[106].EMS[2] AT %DB3810.DBX18950.0, 1 s
   "DB_SDC_EMS_TS_1_HMI_SEK[107].EMS[2]" : UDT_SDC_EMS_TS_STAT_HMI = PLC DB_SDC_EMS_TS_1_HMI.SEK[107].EMS[2] AT %DB3810.DBX19130.0, 1 s
   "DB_SDC_EMS_TS_1_HMI_SEK[108].EMS[2]" : UDT_SDC_EMS_TS_STAT_HMI = PLC DB_SDC_EMS_TS_1_HMI.SEK[108].EMS[2] AT %DB3810.DBX19310.0, 1 s
   "DB_SDC_EMS_TS_1_HMI_SEK[109].EMS[2]" : UDT_SDC_EMS_TS_STAT_HMI = PLC DB_SDC_EMS_TS_1_HMI.SEK[109].EMS[2] AT %DB3810.DBX19490.0, 1 s
   "DB_SDC_EMS_TS_1_HMI_SEK[110].EMS[2]" : UDT_SDC_EMS_TS_STAT_HMI = PLC DB_SDC_EMS_TS_1_HMI.SEK[110].EMS[2] AT %DB3810.DBX19670.0, 1 s
   "DB_SDC_EMS_TS_1_HMI_SEK[111].EMS[2]" : UDT_SDC_EMS_TS_STAT_HMI = PLC DB_SDC_EMS_TS_1_HMI.SEK[111].EMS[2] AT %DB3810.DBX19850.0, 1 s
   "DB_SDC_EMS_TS_1_HMI_SEK[112].EMS[2]" : UDT_SDC_EMS_TS_STAT_HMI = PLC DB_SDC_EMS_TS_1_HMI.SEK[112].EMS[2] AT %DB3810.DBX20030.0, 1 s
   "DB_SDC_EMS_TS_1_HMI_SEK[113].EMS[2]" : UDT_SDC_EMS_TS_STAT_HMI = PLC DB_SDC_TS_PARAMETER_4.HEADER.MAX_NR_SEK AT %DB3810.DBX20210.0, 1 s
   "DB_SDC_EMS_TS_1_HMI_SEK[114].EMS[2]" : UDT_SDC_EMS_TS_STAT_HMI = PLC DB_SDC_EMS_TS_1_HMI.SEK[114].EMS[2] AT %DB3810.DBX20390.0, 1 s
   "DB_SDC_EMS_TS_2_HMI_SEK[204].EMS[1]" : UDT_SDC_EMS_TS_STAT_HMI = PLC DB_SDC_EMS_TS_2_HMI.SEK[204].EMS[1] AT %DB3811.DBX560.0, 1 s
   "DB_SDC_EMS_TS_2_HMI_SEK[204].EMS[2]" : UDT_SDC_EMS_TS_STAT_HMI = PLC DB_SDC_EMS_TS_2_HMI.SEK[204].EMS[2] AT %DB3811.DBX590.0, 1 s
   "DB_SDC_EMS_TS_2_HMI_SEK[205].EMS[1]" : UDT_SDC_EMS_TS_STAT_HMI = PLC DB_SDC_EMS_TS_2_HMI.SEK[205].EMS[1] AT %DB3811.DBX740.0, 1 s
   "DB_SDC_EMS_TS_2_HMI_SEK[205].EMS[2]" : UDT_SDC_EMS_TS_STAT_HMI = PLC DB_SDC_EMS_TS_2_HMI.SEK[205].EMS[2] AT %DB3811.DBX770.0, 1 s
   "DB_SDC_EMS_TS_2_HMI_SEK[206].EMS[1]" : UDT_SDC_EMS_TS_STAT_HMI = PLC DB_SDC_EMS_TS_2_HMI.SEK[206].EMS[1] AT %DB3811.DBX920.0, 1 s
   "DB_SDC_EMS_TS_2_HMI_SEK[206].EMS[2]" : UDT_SDC_EMS_TS_STAT_HMI = PLC DB_SDC_EMS_TS_2_HMI.SEK[206].EMS[2] AT %DB3811.DBX950.0, 1 s
   "DB_SDC_EMS_TS_2_HMI_SEK[207].EMS[1]" : UDT_SDC_EMS_TS_STAT_HMI = PLC DB_SDC_EMS_TS_2_HMI.SEK[207].EMS[1] AT %DB3811.DBX1100.0, 1 s
   "DB_SDC_EMS_TS_2_HMI_SEK[207].EMS[2]" : UDT_SDC_EMS_TS_STAT_HMI = PLC DB_SDC_EMS_TS_2_HMI.SEK[207].EMS[2] AT %DB3811.DBX1130.0, 1 s
   "DB_SDC_EMS_TS_2_HMI_SEK[208].EMS[1]" : UDT_SDC_EMS_TS_STAT_HMI = PLC DB_SDC_EMS_TS_2_HMI.SEK[208].EMS[1] AT %DB3811.DBX1280.0, 1 s
   "DB_SDC_EMS_TS_2_HMI_SEK[208].EMS[2]" : UDT_SDC_EMS_TS_STAT_HMI = PLC DB_SDC_EMS_TS_2_HMI.SEK[208].EMS[2] AT %DB3811.DBX1310.0, 1 s
   "DB_SDC_EMS_TS_2_HMI_SEK[209].EMS[1]" : UDT_SDC_EMS_TS_STAT_HMI = PLC DB_SDC_EMS_TS_2_HMI.SEK[209].EMS[1] AT %DB3811.DBX1460.0, 1 s
   "DB_SDC_EMS_TS_2_HMI_SEK[209].EMS[2]" : UDT_SDC_EMS_TS_STAT_HMI = PLC DB_SDC_EMS_TS_2_HMI.SEK[209].EMS[2] AT %DB3811.DBX1490.0, 1 s
   "DB_SDC_EMS_TS_2_HMI_SEK[210].EMS[1]" : UDT_SDC_EMS_TS_STAT_HMI = PLC DB_SDC_EMS_TS_2_HMI.SEK[210].EMS[1] AT %DB3811.DBX1640.0, 1 s
   "DB_SDC_EMS_TS_2_HMI_SEK[210].EMS[2]" : UDT_SDC_EMS_TS_STAT_HMI = PLC DB_SDC_EMS_TS_2_HMI.SEK[210].EMS[2] AT %DB3811.DBX1670.0, 1 s
   "DB_SDC_EMS_TS_2_HMI_SEK[230].EMS[1]" : UDT_SDC_EMS_TS_STAT_HMI = PLC DB_SDC_EMS_TS_2_HMI.SEK[230].EMS[1] AT %DB3811.DBX5240.0, 1 s
   "DB_SDC_EMS_TS_2_HMI_SEK[230].EMS[2]" : UDT_SDC_EMS_TS_STAT_HMI = PLC DB_SDC_EMS_TS_2_HMI.SEK[230].EMS[2] AT %DB3811.DBX5270.0, 1 s
   "DB_SDC_EMS_TS_2_HMI_SEK[231].EMS[1]" : UDT_SDC_EMS_TS_STAT_HMI = PLC DB_SDC_EMS_TS_2_HMI.SEK[231].EMS[1] AT %DB3811.DBX5420.0, 1 s
   "DB_SDC_EMS_TS_2_HMI_SEK[231].EMS[2]" : UDT_SDC_EMS_TS_STAT_HMI = PLC DB_SDC_EMS_TS_2_HMI.SEK[231].EMS[2] AT %DB3811.DBX5450.0, 1 s
   "DB_SDC_EMS_TS_2_HMI_SEK[232].EMS[1]" : UDT_SDC_EMS_TS_STAT_HMI = PLC DB_SDC_EMS_TS_2_HMI.SEK[232].EMS[1] AT %DB3811.DBX5600.0, 1 s
   "DB_SDC_EMS_TS_2_HMI_SEK[232].EMS[2]" : UDT_SDC_EMS_TS_STAT_HMI = PLC DB_SDC_EMS_TS_2_HMI.SEK[232].EMS[2] AT %DB3811.DBX5630.0, 1 s
   "DB_SDC_EMS_TS_2_HMI_SEK[233].EMS[1]" : UDT_SDC_EMS_TS_STAT_HMI = PLC DB_SDC_EMS_TS_2_HMI.SEK[233].EMS[1] AT %DB3811.DBX5780.0, 1 s
   "DB_SDC_EMS_TS_2_HMI_SEK[233].EMS[2]" : UDT_SDC_EMS_TS_STAT_HMI = PLC DB_SDC_EMS_TS_2_HMI.SEK[233].EMS[2] AT %DB3811.DBX5810.0, 1 s
   "DB_SDC_EMS_TS_2_HMI_SEK[234].EMS[1]" : UDT_SDC_EMS_TS_STAT_HMI = PLC DB_SDC_EMS_TS_2_HMI.SEK[234].EMS[1] AT %DB3811.DBX5960.0, 1 s
   "DB_SDC_EMS_TS_2_HMI_SEK[234].EMS[2]" : UDT_SDC_EMS_TS_STAT_HMI = PLC DB_SDC_EMS_TS_2_HMI.SEK[234].EMS[2] AT %DB3811.DBX5990.0, 1 s
   "DB_SDC_EMS_TS_2_HMI_SEK[235].EMS[1]" : UDT_SDC_EMS_TS_STAT_HMI = PLC DB_SDC_EMS_TS_2_HMI.SEK[235].EMS[1] AT %DB3811.DBX6140.0, 1 s
   "DB_SDC_EMS_TS_2_HMI_SEK[235].EMS[2]" : UDT_SDC_EMS_TS_STAT_HMI = PLC DB_SDC_EMS_TS_2_HMI.SEK[235].EMS[2] AT %DB3811.DBX6170.0, 1 s

